// TIA Portal project "plc_main_V16" (V16)

(* hardware
DEVICE "S7-1200 station_1"  S7-1200 Station
   slot 0: "Rack_0"  S7-1200 Rack  Rack  V1.0
   slot 1: "PLC_main_ip_net_8"  CPU 1215C DC/DC/DC  6ES7 215-1AG40-0XB0  V4.2
DEVICE "PC-System_1"  SIMATIC PC station
   slot 0: "SIMATIC PC station"  Rail  SIMATIC PC-Station  V1.0
      slot 125: "Stationmanager"  Station_Manager  V6.0.4
   slot 1: "HMI_RT_1"  WinCC RT Advanced  6AV2 104-0xxxx-xxxx  16.0.0.0
      slot 33792: "Computer interface"  Host interface
   slot 2: "IE general_1"  IE General  IE_CP  V8.2.0
*)

// ===== PLC "PLC_main_ip_net_8"  CPU 1215C DC/DC/DC =====

VAR_GLOBAL   // PLC tag table "Default tag table"
   "Tag_1" AT %Q0.0 : Bool;
   "Tag_2" AT %Q0.1 : Bool;
   "LOGO_VM2" AT %MB100 : Byte;
   "LOGO_VM2.0" AT %M100.0 : Bool;
END_VAR

// folder: LGF/1 Date and timer operations/LGF_Astro

TYPE "LGF_typeAstroDMS"
VERSION : 0.1
   STRUCT
      dir : Char;   // Direction [N, S, E, W, n, s, e, w]
      deg : UInt;   // Degrees LAT [-89..+ 89]; LON [-179..+179]
      min : UInt;   // Minutes [0..+59]
      sec : UInt;   // Seconds [0..+59]
   END_STRUCT;
END_TYPE

// folder: LGF/8 Technology operations/LGF_NonLin

TYPE "LGF_typeNonLinSetpoints"
VERSION : 0.1
   STRUCT
      InputValue : Real;
      OutputValue : Real;
   END_STRUCT;
END_TYPE

// folder: LGF/8 Technology operations/LGF_Ramp

TYPE "LGF_typeRampTimeTable"
   STRUCT
      outVal : Real;
      "time" : Time;
   END_STRUCT;
END_TYPE

// folder: LGF/9 Measurement operations/LGF_RegressionLine

TYPE "LGF_typeRegressionLine"
   STRUCT
      x : Real;
      y : Real;
   END_STRUCT;
END_TYPE

// folder: Control_functions

DATA_BLOCK "control_DB"   // DB6
{ S7_Optimized_Access := 'FALSE' }
VERSION : 0.1
   VAR
      temperature_setpoint : Int;
      max_presure : Int := 40;
      emerg_coll_down : Bool;
      presure_err : Bool;
   END_VAR
BEGIN
END_DATA_BLOCK

DATA_BLOCK "LOGO"   // DB7
{ S7_Optimized_Access := 'FALSE' }
VERSION : 0.1
   VAR
      LOGO_heating_state : Bool;
   END_VAR
BEGIN
END_DATA_BLOCK

DATA_BLOCK "sensor_inputs"   // DB8
{ S7_Optimized_Access := 'TRUE' }
VERSION : 0.1
   VAR
      burning_temperature : Int;
      fire_state : Bool;
      flow_speed : Int;
      fluid_t : Int;
      system_presure : Int;
   END_VAR
BEGIN
END_DATA_BLOCK

DATA_BLOCK "actuators_output"   // DB9
{ S7_Optimized_Access := 'FALSE' }
VERSION : 0.1
   VAR
      gas_flow : Int;
      pimp_speed : Int;
      valve_state : Bool;
   END_VAR
BEGIN
END_DATA_BLOCK

DATA_BLOCK "Main_control_DB"   // DB10
{ S7_Optimized_Access := 'TRUE' }
VERSION : 0.1
// stored: InstanceOfName Main_control
"Main_control"
BEGIN
END_DATA_BLOCK

DATA_BLOCK "LGF_Impulse_DB_2"   // DB11
{ S7_Optimized_Access := 'TRUE' }
VERSION : 0.1
// stored: InstanceOfName LGF_Impulse
"LGF_Impulse"
BEGIN
END_DATA_BLOCK

// folder: Phisical_functions

DATA_BLOCK "phisical_DB"   // DB1
{ S7_Optimized_Access := 'TRUE' }
VERSION : 0.1
   VAR
      burning_t_old : Int;
      OUT_burning_t : Int;
      OUT_fire_state : Bool;
      OUT_fluid_t : Int;
      OUT_flow_speed : Int;
      IN_gas_flow : Int;
      IN_pimp_speed : Int;
      IN_valve_state : Bool;
      IN_pump_state : Bool;
      OUT_pump_err : Bool;
      OUT_pipe_err : Bool;
      OUT_tank_err : Bool;
      OUT_tank_presure : Int;
      OUT_residential_heeting : Bool;
      pump_failure : Bool := false;
      tank_failure : Bool := false;
      max_pump_failure_time : Time := T#10s;
      max_tank_presure : Int := 50;
   END_VAR
BEGIN
END_DATA_BLOCK

DATA_BLOCK "LGF_Impulse_DB"   // DB2
{ S7_Optimized_Access := 'TRUE' }
VERSION : 0.1
// stored: InstanceOfName LGF_Impulse
"LGF_Impulse"
BEGIN
END_DATA_BLOCK

DATA_BLOCK "LGF_Impulse_DB_1"   // DB3
{ S7_Optimized_Access := 'TRUE' }
VERSION : 0.1
// stored: InstanceOfName LGF_Impulse
"LGF_Impulse"
BEGIN
END_DATA_BLOCK

DATA_BLOCK "Phisical_proces_sim_dont_touch_DB_1"   // DB4
{ S7_Optimized_Access := 'TRUE' }
VERSION : 0.1
// stored: InstanceOfName Phisical_proces_sim_dont_touch
"Phisical_proces_sim_dont_touch"
BEGIN
END_DATA_BLOCK

// folder: System blocks/Program resources

DATA_BLOCK "IEC_Timer_0_DB"   // DB5
{ S7_Optimized_Access := 'TRUE' }
AUTHOR : Simatic
FAMILY : IEC
NAME : IEC_TMR
VERSION : 1.0
// stored: InstanceOfName IEC_TIMER
"IEC_TIMER"
BEGIN
END_DATA_BLOCK

// folder: (top level)

ORGANIZATION_BLOCK "Main"   // OB1, LAD, ProgramCycle
TITLE = "Main Program Sweep (Cycle)"
{ S7_Optimized_Access := 'TRUE' }
VERSION : 0.1
   VAR_INPUT
      Initial_Call : Bool;   // Initial call of this OB
      Remanence : Bool;   // =True, if remanent data are available
   END_VAR
BEGIN

REGION Network 1: Phisical proces
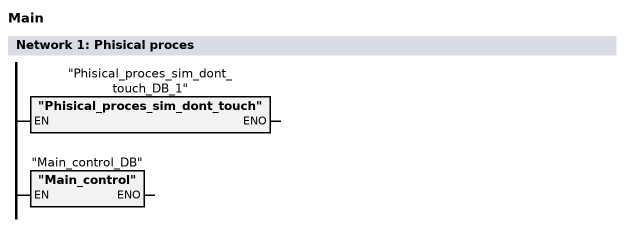
   RUNG wire#powerrail
      "Phisical_proces_sim_dont_touch_DB_1"()
   END_RUNG
   RUNG wire#powerrail
      "Main_control_DB"()
   END_RUNG
   // the same network as SCL:
   "Phisical_proces_sim_dont_touch_DB_1"();   // "Phisical_proces_sim_dont_touch"
   "Main_control_DB"();   // "Main_control"
END_REGION
END_ORGANIZATION_BLOCK

// folder: Control_functions

FUNCTION_BLOCK "Main_control"   // FB6, LAD
{ S7_Optimized_Access := 'TRUE' }
VERSION : 0.1
BEGIN

REGION Network 1
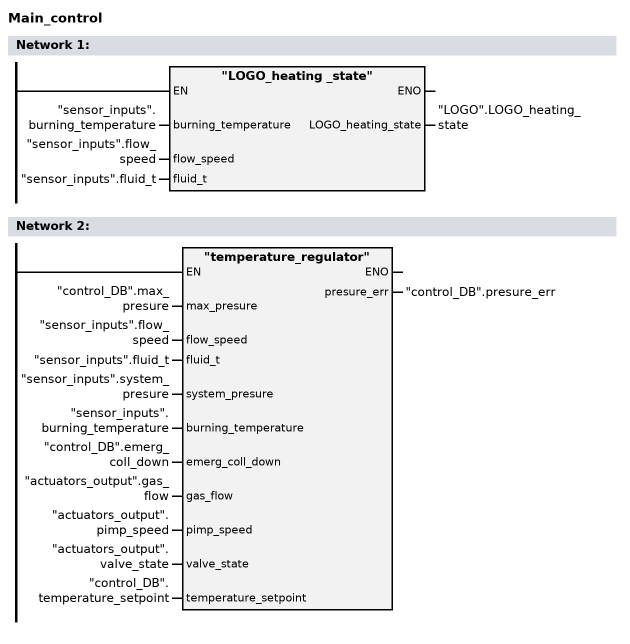
   RUNG wire#powerrail
      "LOGO_heating _state"(burning_temperature := "sensor_inputs".burning_temperature, flow_speed := "sensor_inputs".flow_speed, fluid_t := "sensor_inputs".fluid_t, LOGO_heating_state => "LOGO".LOGO_heating_state)
   END_RUNG
   // the same network as SCL:
   "LOGO_heating _state"(burning_temperature := "sensor_inputs".burning_temperature,
                         flow_speed := "sensor_inputs".flow_speed,
                         fluid_t := "sensor_inputs".fluid_t,
                         LOGO_heating_state => "LOGO".LOGO_heating_state);
END_REGION

REGION Network 2
   RUNG wire#powerrail
      "temperature_regulator"(max_presure := "control_DB".max_presure, flow_speed := "sensor_inputs".flow_speed, fluid_t := "sensor_inputs".fluid_t, system_presure := "sensor_inputs".system_presure, burning_temperature := "sensor_inputs".burning_temperature, emerg_coll_down := "control_DB".emerg_coll_down, gas_flow := "actuators_output".gas_flow, pimp_speed := "actuators_output".pimp_speed, valve_state := "actuators_output".valve_state, temperature_setpoint := "control_DB".temperature_setpoint, presure_err => "control_DB".presure_err)
   END_RUNG
   // the same network as SCL:
   "temperature_regulator"(max_presure := "control_DB".max_presure,
                           flow_speed := "sensor_inputs".flow_speed,
                           fluid_t := "sensor_inputs".fluid_t,
                           system_presure := "sensor_inputs".system_presure,
                           burning_temperature := "sensor_inputs".burning_temperature,
                           emerg_coll_down := "control_DB".emerg_coll_down,
                           gas_flow := "actuators_output".gas_flow,
                           pimp_speed := "actuators_output".pimp_speed,
                           valve_state := "actuators_output".valve_state,
                           temperature_setpoint := "control_DB".temperature_setpoint,
                           presure_err => "control_DB".presure_err);
END_REGION
END_FUNCTION_BLOCK

FUNCTION "LOGO_heating _state" : Void   // FC12, SCL
{ S7_Optimized_Access := 'TRUE' }
VERSION : 0.1
   VAR_INPUT
      burning_temperature : Int;
      flow_speed : Int;
      fluid_t : Int;
   END_VAR
   VAR_OUTPUT
      LOGO_heating_state : Bool;
   END_VAR
BEGIN
   IF #flow_speed > 1 AND #fluid_t > 15 THEN
       // Statement section IF
       #LOGO_heating_state := TRUE;
   ELSE
       #LOGO_heating_state := FALSE;
   END_IF;
END_FUNCTION

FUNCTION "temperature_regulator" : Void   // FC15, SCL
{ S7_Optimized_Access := 'TRUE' }
VERSION : 0.1
   VAR_INPUT
      max_presure : Int;
      flow_speed : Int;
      fluid_t : Int;
      system_presure : Int;
      burning_temperature : Int;
   END_VAR
   VAR_OUTPUT
      presure_err : Bool;
   END_VAR
   VAR_IN_OUT
      emerg_coll_down : Bool;
      gas_flow : Int;
      pimp_speed : Int;
      valve_state : Bool;
      temperature_setpoint : Int;
   END_VAR
   VAR_TEMP
      impulse : Bool;
   END_VAR
BEGIN
   "LGF_Impulse_DB_2"(frequency:=0.7,
                      impulse=>#impulse);

   IF #system_presure > #max_presure THEN
       // Statement section IF
       #temperature_setpoint := 0;
       #presure_err := true;
   END_IF;

   IF #impulse = TRUE THEN
       IF #temperature_setpoint > 0 THEN
           // Statement section IF
           #pimp_speed := 869;
       ELSE
           IF #pimp_speed > 0 THEN
               // Statement section IF
               #pimp_speed := #pimp_speed - 1;
           ELSE
               #pimp_speed := 0;
           END_IF;


       END_IF;
       // Statement section IF
       IF #temperature_setpoint > #fluid_t THEN
           // Statement section IF
           #gas_flow := #gas_flow + 1;
       ELSIF #temperature_setpoint < #fluid_t THEN
           #gas_flow := #gas_flow - 1;
       END_IF;

   END_IF;
END_FUNCTION

// folder: Phisical_functions

FUNCTION_BLOCK "Phisical_proces_sim_dont_touch"   // FB1, LAD
{ S7_Optimized_Access := 'TRUE' }
VERSION : 0.1
BEGIN

REGION Network 1
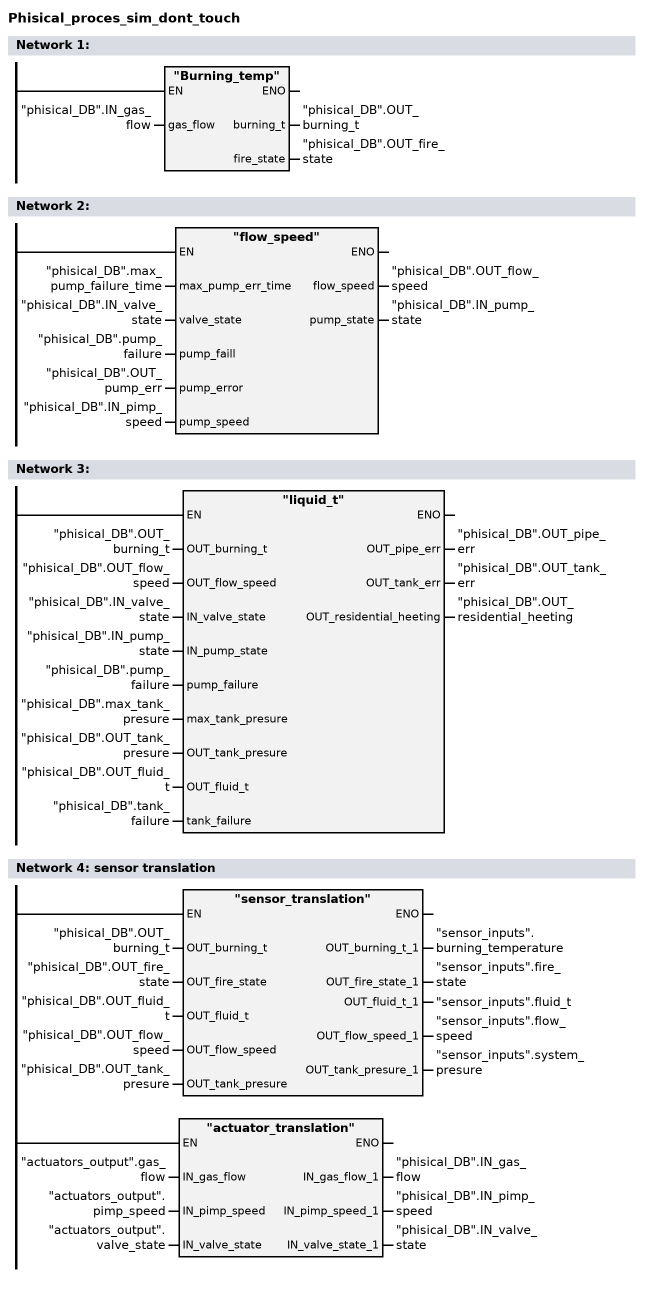
   RUNG wire#powerrail
      "Burning_temp"(gas_flow := "phisical_DB".IN_gas_flow, burning_t => "phisical_DB".OUT_burning_t, fire_state => "phisical_DB".OUT_fire_state)
   END_RUNG
   // the same network as SCL:
   "Burning_temp"(gas_flow := "phisical_DB".IN_gas_flow,
                  burning_t => "phisical_DB".OUT_burning_t,
                  fire_state => "phisical_DB".OUT_fire_state);
END_REGION

REGION Network 2
   RUNG wire#powerrail
      "flow_speed"(max_pump_err_time := "phisical_DB".max_pump_failure_time, valve_state := "phisical_DB".IN_valve_state, pump_faill := "phisical_DB".pump_failure, pump_error := "phisical_DB".OUT_pump_err, pump_speed := "phisical_DB".IN_pimp_speed, flow_speed => "phisical_DB".OUT_flow_speed, pump_state => "phisical_DB".IN_pump_state)
   END_RUNG
   // the same network as SCL:
   "flow_speed"(max_pump_err_time := "phisical_DB".max_pump_failure_time,
                valve_state := "phisical_DB".IN_valve_state,
                pump_faill := "phisical_DB".pump_failure,
                pump_error := "phisical_DB".OUT_pump_err,
                pump_speed := "phisical_DB".IN_pimp_speed,
                flow_speed => "phisical_DB".OUT_flow_speed,
                pump_state => "phisical_DB".IN_pump_state);
END_REGION

REGION Network 3
   RUNG wire#powerrail
      "liquid_t"(OUT_burning_t := "phisical_DB".OUT_burning_t, OUT_flow_speed := "phisical_DB".OUT_flow_speed, IN_valve_state := "phisical_DB".IN_valve_state, IN_pump_state := "phisical_DB".IN_pump_state, pump_failure := "phisical_DB".pump_failure, max_tank_presure := "phisical_DB".max_tank_presure, OUT_tank_presure := "phisical_DB".OUT_tank_presure, OUT_fluid_t := "phisical_DB".OUT_fluid_t, tank_failure := "phisical_DB".tank_failure, OUT_pipe_err => "phisical_DB".OUT_pipe_err, OUT_tank_err => "phisical_DB".OUT_tank_err, OUT_residential_heeting => "phisical_DB".OUT_residential_heeting)
   END_RUNG
   // the same network as SCL:
   "liquid_t"(OUT_burning_t := "phisical_DB".OUT_burning_t,
              OUT_flow_speed := "phisical_DB".OUT_flow_speed,
              IN_valve_state := "phisical_DB".IN_valve_state,
              IN_pump_state := "phisical_DB".IN_pump_state,
              pump_failure := "phisical_DB".pump_failure,
              max_tank_presure := "phisical_DB".max_tank_presure,
              OUT_tank_presure := "phisical_DB".OUT_tank_presure,
              OUT_fluid_t := "phisical_DB".OUT_fluid_t,
              tank_failure := "phisical_DB".tank_failure,
              OUT_pipe_err => "phisical_DB".OUT_pipe_err,
              OUT_tank_err => "phisical_DB".OUT_tank_err,
              OUT_residential_heeting => "phisical_DB".OUT_residential_heeting);
END_REGION

REGION Network 4: sensor translation
   RUNG wire#powerrail
      "sensor_translation"(OUT_burning_t := "phisical_DB".OUT_burning_t, OUT_fire_state := "phisical_DB".OUT_fire_state, OUT_fluid_t := "phisical_DB".OUT_fluid_t, OUT_flow_speed := "phisical_DB".OUT_flow_speed, OUT_tank_presure := "phisical_DB".OUT_tank_presure, OUT_burning_t_1 => "sensor_inputs".burning_temperature, OUT_fire_state_1 => "sensor_inputs".fire_state, OUT_fluid_t_1 => "sensor_inputs".fluid_t, OUT_flow_speed_1 => "sensor_inputs".flow_speed, OUT_tank_presure_1 => "sensor_inputs".system_presure)
   END_RUNG
   RUNG wire#powerrail
      "actuator_translation"(IN_gas_flow := "actuators_output".gas_flow, IN_pimp_speed := "actuators_output".pimp_speed, IN_valve_state := "actuators_output".valve_state, IN_gas_flow_1 => "phisical_DB".IN_gas_flow, IN_pimp_speed_1 => "phisical_DB".IN_pimp_speed, IN_valve_state_1 => "phisical_DB".IN_valve_state)
   END_RUNG
   // the same network as SCL:
   "sensor_translation"(OUT_burning_t := "phisical_DB".OUT_burning_t,
                        OUT_fire_state := "phisical_DB".OUT_fire_state,
                        OUT_fluid_t := "phisical_DB".OUT_fluid_t,
                        OUT_flow_speed := "phisical_DB".OUT_flow_speed,
                        OUT_tank_presure := "phisical_DB".OUT_tank_presure,
                        OUT_burning_t_1 => "sensor_inputs".burning_temperature,
                        OUT_fire_state_1 => "sensor_inputs".fire_state,
                        OUT_fluid_t_1 => "sensor_inputs".fluid_t,
                        OUT_flow_speed_1 => "sensor_inputs".flow_speed,
                        OUT_tank_presure_1 => "sensor_inputs".system_presure);
   "actuator_translation"(IN_gas_flow := "actuators_output".gas_flow,
                          IN_pimp_speed := "actuators_output".pimp_speed,
                          IN_valve_state := "actuators_output".valve_state,
                          IN_gas_flow_1 => "phisical_DB".IN_gas_flow,
                          IN_pimp_speed_1 => "phisical_DB".IN_pimp_speed,
                          IN_valve_state_1 => "phisical_DB".IN_valve_state);
END_REGION
END_FUNCTION_BLOCK

FUNCTION "Burning_temp" : Void   // FC1, SCL
{ S7_Optimized_Access := 'TRUE' }
VERSION : 0.1
   VAR_INPUT
      gas_flow : Int;
   END_VAR
   VAR_OUTPUT
      burning_t : Int;
      fire_state : Bool;
   END_VAR
   VAR_TEMP
      burning_t_temp : Int;
      triger : Bool;
   END_VAR
   VAR CONSTANT
      gas_to_temp : Int := 2;
   END_VAR
BEGIN
   //generates gas input state based on gas flow
   IF #gas_flow = 0 THEN
       #fire_state := FALSE;
   ELSE
       #fire_state := TRUE;
   END_IF;

   //Writing to phisicalDB
   #burning_t := #gas_flow * #gas_to_temp;
END_FUNCTION

FUNCTION "flow_speed" : Void   // FC10, SCL
{ S7_Optimized_Access := 'TRUE' }
VERSION : 0.1
   VAR_INPUT
      max_pump_err_time : Time;
      valve_state : Bool;
   END_VAR
   VAR_OUTPUT
      flow_speed : Int;
      pump_state : Bool;
   END_VAR
   VAR_IN_OUT
      pump_faill : Bool;
      pump_error : Bool;
      pump_speed : Int;
   END_VAR
   VAR_TEMP
      pump_err : Bool;
      impulse : Bool;
      countdown : Time;
      fault_timer_reset : Bool;
   END_VAR
   VAR CONSTANT
      rpm_to_l : Int := 10;
   END_VAR
BEGIN

   "LGF_Impulse_DB_1"(frequency:=70.0,
                      impulse=>#impulse,
                      countdown=>#countdown);

   IF #pump_faill = FALSE THEN
       // Statement section IF
       IF #pump_speed = 0 THEN
           // Statement section IF
           #pump_state := FALSE;
           #pump_err := FALSE;
       ELSE
           #pump_state := TRUE;

           IF #valve_state = FALSE THEN
               #flow_speed := 0;
               #pump_err := TRUE;
           ELSE

               #flow_speed := #pump_speed / #rpm_to_l;
               #pump_err := FALSE;

           END_IF;

       END_IF;
   ELSE
       #pump_state := TRUE;
       #pump_err := TRUE;
       #flow_speed := 0;
   END_IF;



       #pump_error := #pump_err;

       IF #pump_error = FALSE AND #pump_faill = FALSE THEN
           #fault_timer_reset := TRUE;
       ELSE
           #fault_timer_reset := FALSE;
       END_IF;

       "IEC_Timer_0_DB".TONR(IN:=#pump_error,
                             R:=#fault_timer_reset,
                             PT:=#max_pump_err_time,
                             Q=>#pump_faill
       );
END_FUNCTION

FUNCTION "liquid_t" : Void   // FC11, SCL
{ S7_Optimized_Access := 'TRUE' }
VERSION : 0.1
   VAR_INPUT
      OUT_burning_t : Int;
      OUT_flow_speed : Int;
      IN_valve_state : Bool;
      IN_pump_state : Bool;
      pump_failure : Bool;
      max_tank_presure : Int;
   END_VAR
   VAR_OUTPUT
      OUT_pipe_err : Bool;
      OUT_tank_err : Bool;
      OUT_residential_heeting : Bool;
   END_VAR
   VAR_IN_OUT
      OUT_tank_presure : Int;
      OUT_fluid_t : Int;
      tank_failure : Bool;
   END_VAR
   VAR_TEMP
      impulse : Bool;
      countdown : Time;
      valv_closes_increase : Int;
      pump_heat_decrease : Int;
      fluid_calculated_current : Int;
   END_VAR
   VAR CONSTANT
      fluid_to_burning_ratio : Int := 3;
   END_VAR
BEGIN
   "LGF_Impulse_DB"(frequency:=1.0,
                    impulse=>#impulse,
                    countdown=>#countdown);

   #valv_closes_increase := 0;

   #fluid_calculated_current := (#OUT_burning_t / #fluid_to_burning_ratio);

   (* IF #IN_valve_state = TRUE AND #IN_pump_state = TRUE THEN
       // Statement section IF
       #fluid_calculated_current := #fluid_calculated_current - #OUT_flow_speed / 8;
   END_IF; *)

   IF #impulse THEN


       (*
       HOW to create it so that when pump and valve doesnt work, temperature slowly increases
       *)

       IF #IN_valve_state = FALSE OR #IN_pump_state = FALSE OR #pump_failure = TRUE THEN

           IF #OUT_burning_t > #OUT_fluid_t THEN
               // Statement section IF
               #OUT_fluid_t := #OUT_fluid_t + 1;
           END_IF;

           IF #OUT_burning_t < #OUT_fluid_t THEN
               // Statement section IF
               #OUT_fluid_t := #OUT_fluid_t - 1;
           END_IF;

       ELSE
           IF #fluid_calculated_current > #OUT_fluid_t THEN
               // Statement section IF
               #OUT_fluid_t := #OUT_fluid_t + 1;
           END_IF;

           IF #fluid_calculated_current < #OUT_fluid_t THEN
               // Statement section IF
               #OUT_fluid_t := #OUT_fluid_t - 1;
           END_IF;
       END_IF;

       IF #tank_failure = TRUE THEN
           // Statement section IF
           #OUT_tank_presure := #OUT_tank_presure - 5;
       ELSE
           #OUT_tank_presure := ((#OUT_fluid_t) / 2.83);
       END_IF;
   END_IF;





   IF #tank_failure = FALSE THEN
       IF #OUT_tank_presure > #max_tank_presure THEN
           #tank_failure := TRUE;
       END_IF;
   END_IF;



   IF #OUT_fluid_t > 30 & #IN_valve_state = TRUE & #IN_pump_state = TRUE THEN
       IF #pump_failure = TRUE THEN

           #OUT_residential_heeting := FALSE;
       ELSE
           #OUT_residential_heeting := TRUE;
       END_IF;


   ELSE
       #OUT_residential_heeting := FALSE;
   END_IF;
END_FUNCTION

FUNCTION "sensor_translation" : Void   // FC13, SCL
{ S7_Optimized_Access := 'TRUE' }
VERSION : 0.1
   VAR_INPUT
      OUT_burning_t : Int;
      OUT_fire_state : Bool;
      OUT_fluid_t : Int;
      OUT_flow_speed : Int;
      OUT_tank_presure : Int;
   END_VAR
   VAR_OUTPUT
      OUT_burning_t_1 : Int;
      OUT_fire_state_1 : Bool;
      OUT_fluid_t_1 : Int;
      OUT_flow_speed_1 : Int;
      OUT_tank_presure_1 : Int;
   END_VAR
BEGIN
   #OUT_burning_t_1 := #OUT_burning_t;
   #OUT_fire_state_1 := #OUT_fire_state;
   #OUT_fluid_t_1 := #OUT_fluid_t;
   #OUT_flow_speed_1 := #OUT_flow_speed;
   #OUT_tank_presure_1 := #OUT_tank_presure;
END_FUNCTION

FUNCTION "actuator_translation" : Void   // FC14, SCL
{ S7_Optimized_Access := 'TRUE' }
VERSION : 0.1
   VAR_INPUT
      IN_gas_flow : Int;
      IN_pimp_speed : Int;
      IN_valve_state : Bool;
   END_VAR
   VAR_OUTPUT
      IN_gas_flow_1 : Int;
      IN_pimp_speed_1 : Int;
      IN_valve_state_1 : Bool;
   END_VAR
BEGIN
   #IN_gas_flow_1 := #IN_gas_flow;
   #IN_pimp_speed_1 := #IN_pimp_speed;
   #IN_valve_state_1 := #IN_valve_state;
END_FUNCTION

// folder: Phisical_functions/LGF/0 Bit logic operations

FUNCTION_BLOCK "LGF_PulseRelay"   // FB3, SCL
{ S7_Optimized_Access := 'TRUE' }
VERSION : 0.1
   VAR_INPUT
      trigger : Bool;   // trigger signal, rising edge
      set : Bool;   // set signal. rising edge
      reset : Bool;   // reset signal, rising edge
   END_VAR
   VAR_OUTPUT
      out : Bool;   // output signal
   END_VAR
   VAR
      statTriggerOld : Bool := false;   // -
      statTriggerRis : Bool := false;   // -
      statSetOld : Bool := false;   // -
      statSetRis : Bool := false;   // -
      statResetOld : Bool := false;   // -
      statResetRis : Bool := false;   // -
      statOut : Bool := false;   // -
   END_VAR
BEGIN
   //=============================================================================
   // SIEMENS AG
   // (c)Copyright 2017 
   //-----------------------------------------------------------------------------
   // Library:       LGF (Library General Functions)
   // Tested with:   CPU1212C DC/DC/DC FW:V4.2
   // Engineering:   TIA Portal V14 Update 1
   // Restrictions:  -
   // Requirements:  PLC (S7-1200 / S7-1500)
   // Functionality: Pulse relay, Surge relay, Toggle-Flip-Flop, Frequency divider
   //-----------------------------------------------------------------------------
   // Change log table:
   // Version Date        In charge / Changes applied
   // 01.00.00 06.06.2015 Siemens Industry Online Support
   //                     First released version
   // 01.00.01 02.01.2017 Siemens Industry Online Support
   //                     Upgrade: TIA V14 Update 1
   // 01.00.02 02.01.2017 Siemens Industry Online Support
   //                     Comment correction                  
   // 01.00.03 17.08.2018 Siemens Industry Online Support
   //                     Upgrade: TIA V15 Update 2
   // 01.00.04 23.11.2018 Siemens Industry Online Support
   //                     Upgrade: TIA V15.1
   //=============================================================================

   // Scan for risign edge "trigger"
   IF #trigger AND  NOT #statTriggerOld THEN
     #statTriggerRis := TRUE;
   ELSE
     #statTriggerRis := FALSE;
   END_IF;
   #statTriggerOld := #trigger;

   // Scan for risign edge "set"
   IF #set AND NOT #statSetOld THEN
     #statSetRis := TRUE;
   ELSE
     #statSetRis := FALSE;
   END_IF;
   #statSetOld := #set;

   // Scan for risign edge "reset"
   IF #reset AND NOT #statResetOld THEN
     #statResetRis := TRUE;
   ELSE
     #statResetRis := FALSE;
   END_IF;
   #statResetOld := #reset;

   // Create toggle signal
   IF #statTriggerRis AND NOT #statOut THEN
     #statOut := TRUE;
   ELSIF #statTriggerRis AND #statOut THEN
     #statOut := FALSE;
   END_IF;

   // Output: toggle, set, reset
   IF #statTriggerRis THEN
     #out := #statOut;
   END_IF;

   IF #statSetRis THEN
     #out := TRUE;
   END_IF;

   IF #statResetRis THEN
     #out := FALSE;
   END_IF;
END_FUNCTION_BLOCK

// folder: Phisical_functions/LGF/1 Date and timer operations

FUNCTION_BLOCK "LGF_SetTime"   // FB4, SCL
{ S7_Optimized_Access := 'TRUE' }
VERSION : 0.1
   VAR_INPUT
      setSystemTimeUTC : Bool;   // Set system time
      systemTimeUTC : DTL;   // System time
      setLocalTime : Bool;   // Set local time
      localTime : DTL;   // Local Time
      setTimeZone : Bool;   // Set time zone and daylight saving time
      timeZone : Int;   // Timezones HHMM [-1200.. -330.. 0.. 930.. 1200.. 1300]
      daylightSavingTime : Bool;   // Daylight saving time: activated [1], deactivated [0]
   END_VAR
   VAR_OUTPUT
      actSystemTime : DTL;   // -
      actLocalTime : DTL;   // -
      lastSetTimeZone : String;   // Time zone that was set last by this block
      error : Bool;   // Error
      status : Word;   // Status and error codes
      statusID : UInt;   // Error destination: "1" = LGF_SetTime; "2" = SET_TIMEZONE
   END_VAR
   VAR
      statSetSystemTimeOld : Bool;   // -
      statSetLocalTimeOld : Bool;   // -
      statSetTimeZoneOld : Bool;   // -
      statTimeZone : TimeTransformationRule;   // -
      InstSET_TIMEZONE : SET_TIMEZONE;   // -
   END_VAR
   VAR_TEMP
      tempSetLocalTimeRet : Int;   // -
      tempSetSystemTimeRet : Int;   // -
      tempSystemTimeRet : Int;   // -
      tempLocalTimeRet : Int;   // -
      tempTimeZoneDone : Bool;   // -
      tempTimeZoneBusy : Bool;   // -
      tempTimeZoneError : Bool;   // -
      tempTimeZoneStatus : Word;   // -
   END_VAR
   VAR CONSTANT
      HOUR : Int := 60;   // -
      "30MIN" : Int := 30;   // -
      "15MIN" : Int := 15;   // -
      "0MIN" : Int := 0;   // -
      NO_ERROR : Word := 16#0000;   // -
      NO_CURRENT_JOBS : Word := 16#7000;   // -
      ERROR_NO_DEFINED_TIME_ZONE : Word := 16#8200;   // No defined time zone is selected; check input "timeZone"
      ERROR_IN_THIS_BLOCK : UInt := 1;   // Error in this block
      ERROR_SET_TIMEZONE : UInt := 2;   // Error instruction SET_TIMEZONE
   END_VAR
   // statTimeZone.Bias := 0;
   // statTimeZone.DaylightBias := 60;
   // statTimeZone.DaylightStartMonth := 3;
   // statTimeZone.DaylightStartWeek := 5;
   // statTimeZone.DaylightStartWeekday := 1;
   // statTimeZone.DaylightStartHour := 2;
   // statTimeZone.DaylightStartMinute := 0;
   // statTimeZone.StandardStartMonth := 10;
   // statTimeZone.StandardStartWeek := 5;
   // statTimeZone.StandardStartWeekday := 1;
   // statTimeZone.StandardStartHour := 3;
   // statTimeZone.StandardStartMinute := 0;
   // statTimeZone.TimeZoneName := 'not even set by LGF_TimeZone';
BEGIN
   //=============================================================================
   // SIEMENS AG
   // (c)Copyright 2017 
   //-----------------------------------------------------------------------------
   // Library:       LGF (Library General Functions)
   // Tested with:   CPU1212C DC/DC/DC FW:V4.2
   // Engineering:   TIA Portal V14 Update 1
   // Restrictions:  -
   // Requirements:  PLC (S7-1200 / S7-1500)
   // Functionality: Set system time, local time, time zone
   //-----------------------------------------------------------------------------
   // Change log table:
   // Version Date         In charge / Changes applied
   // 01.00.00 08.06.2015  Siemens Industry Online Support
   //                      First released version
   // 01.00.01 02.01.2017  Siemens Industry Online Support
   //                      Upgrade: TIA V14 Update 1
   // 01.00.02 02.03.2017  Siemens Industry Online Support
   //                      Bugfix: FB number: automatic
   // 01.00.03 17.08.2018  Siemens Industry Online Support
   //                      Upgrade: TIA V15 Update 2
   // 01.00.04 23.11.2018  Siemens Industry Online Support
   //                      Upgrade: TIA V15.1
   // 01.00.05 20.02.2019  Siemens Industry Online Support
   //                      Bugfix: Rising edge at input REQ of SET_TIMEOUT
   // =============================================================================

   // Set "No current job" status
   #error := false;
   #statusID := #ERROR_IN_THIS_BLOCK;
   #status := #NO_CURRENT_JOBS;

   // Reading system and local time
   #tempSystemTimeRet := RD_SYS_T(#actSystemTime); // Output current system time
   #tempLocalTimeRet := RD_LOC_T(#actLocalTime); // Output current local

   // Set system time by rising edge =============================================
   IF #setSystemTimeUTC AND NOT #statSetSystemTimeOld THEN
     #tempSetSystemTimeRet := WR_SYS_T(#systemTimeUTC);
   END_IF;
   #statSetSystemTimeOld := #setSystemTimeUTC;

   // Set local time zone by rising edge =========================================
   IF #setLocalTime AND NOT #statSetLocalTimeOld THEN
     #tempSetLocalTimeRet := WR_LOC_T(LOCTIME := #localTime, DST := #daylightSavingTime);
   END_IF;
   #statSetLocalTimeOld := #setLocalTime;

   // Set time zone by rising edge ===============================================
   IF #setTimeZone AND NOT #statSetTimeZoneOld THEN
     CASE #timeZone OF
       -1200:  // (UTC -12:00) Eniwetok, Kwajalein
         #statTimeZone.Bias := -12 * #HOUR;
         #statTimeZone.TimeZoneName := '(UTC -12:00)';
       -1100:  // (UTC -11:00) Midway Island
         #statTimeZone.Bias := -11 * #HOUR;
         #statTimeZone.TimeZoneName := '(UTC -11:00)';
       -1000:  // (UTC -10:00) Hawaii
         #statTimeZone.Bias := -10 * #HOUR;
         #statTimeZone.TimeZoneName := '(UTC -10:00)';
       -930:  // (UTC -09:30) (French) Polynesia
         #statTimeZone.Bias := -9 * #HOUR + #"30MIN";
         #statTimeZone.TimeZoneName := '(UTC -09:00)';
       -900:  // (UTC -09:00) Alaska
         #statTimeZone.Bias := -9 * #HOUR;
         #statTimeZone.TimeZoneName := '(UTC -09:00)';
       -800:  // (UTC -08:00) Tijuana, Los Angeles, Seattle, Vancouver
         #statTimeZone.Bias := -8 * #HOUR;
         #statTimeZone.TimeZoneName := '(UTC -08:00)';
       -700:  // (UTC -07:00) Arizona, Denver, Salt Lake City, Calgary
         #statTimeZone.Bias := -7 * #HOUR;
         #statTimeZone.TimeZoneName := '(UTC -07:00)';
       -600:  // (UTC -06:00) Chicago, Dallas, Kansas City, Winnipeg
         #statTimeZone.Bias := -6 * #HOUR;
         #statTimeZone.TimeZoneName := '(UTC -06:00)';
       -500:  // (UTC -05:00) Eastern Time (USA & Canada)
         #statTimeZone.Bias := -5 * #HOUR;
         #statTimeZone.TimeZoneName := '(UTC -05:00)';
       -400:  // (UTC -04:00) La Paz, Georgetown
         #statTimeZone.Bias := -4 * #HOUR;
         #statTimeZone.TimeZoneName := '(UTC -04:00)';
       -330:  // (UTC -03:30) Newfoundland
         #statTimeZone.Bias := -3 * #HOUR + #"30MIN";
         #statTimeZone.TimeZoneName := '(UTC -03:30)';
       -300:  // (UTC -03:00) Brasilia, Buenos Aires
         #statTimeZone.Bias := -3 * #HOUR;
         #statTimeZone.TimeZoneName := '(UTC -03:00)';
       -200:  // (UTC -02:00) Mid-Atlantic
         #statTimeZone.Bias := -2 * #HOUR;
         #statTimeZone.TimeZoneName := '(UTC -02:00)';
       -100:  // (UTC -01:00) Azores, Cape Verde Is.
         #statTimeZone.Bias := -1 * #HOUR;
         #statTimeZone.TimeZoneName := '(UTC -01:00)';
       0:  // (UTC) Dublin, Edinburgh, Lisbon, London
         #statTimeZone.Bias := 0;
         #statTimeZone.TimeZoneName := '(UTC)';
       100:  // (UTC +01:00) Berlin, Bern, Brussels, Rome, Stockholm, Vienna
         #statTimeZone.Bias := 1 * #HOUR;
         #statTimeZone.TimeZoneName := '(UTC +01:00)';
       200: // (UTC +02:00) Athens, Istanbul, Minsk, Bucharest
         #statTimeZone.Bias := 2 * #HOUR;
         #statTimeZone.TimeZoneName := '(UTC +02:00)';
       300: // (UTC +03:00) Baghdad, Kuwait, Riyadh
         #statTimeZone.Bias := 3 * #HOUR;
         #statTimeZone.TimeZoneName := '(UTC +03:00)';
       330: // (UTC +03:00) Iran
         #statTimeZone.Bias := 3 * #HOUR + #"30MIN";
         #statTimeZone.TimeZoneName := '(UTC +03:30)';
       400: // (UTC +04:00) Moscow, St. Petersburg, Volgograd, Abu Dhabi, Muscat
         #statTimeZone.Bias := 4 * #HOUR;
         #statTimeZone.TimeZoneName := '(UTC +04:00)';
       430: // (UTC +04:30) Afghanistan
         #statTimeZone.Bias := 4 * #HOUR + #"30MIN";
         #statTimeZone.TimeZoneName := '(UTC +04:30)';
       500: // (UTC +05:00) Islamabad, Karachi, Tashkent
         #statTimeZone.Bias := 5 * #HOUR;
         #statTimeZone.TimeZoneName := '(UTC +05:00)';
       530: // (UTC +05:30) India, Sri Lanka
         #statTimeZone.Bias := 5 * #HOUR + #"30MIN";
         #statTimeZone.TimeZoneName := '(UTC +05:30)';
       545: // (UTC +05:45) India, Sri Lanka
         #statTimeZone.Bias := 5 * #HOUR + #"30MIN" + #"15MIN";
         #statTimeZone.TimeZoneName := '(UTC +05:45)';
       600: // (UTC +06:00) Astana, Almaty, Dhaka, Colombo
         #statTimeZone.Bias := 6 * #HOUR;
         #statTimeZone.TimeZoneName := '(UTC +06:00)';
       630: // (UTC +06:30) Coco Island, Mayanmar
         #statTimeZone.Bias := 6 * #HOUR + #"30MIN";
         #statTimeZone.TimeZoneName := '(UTC +06:30)';
       700: // (UTC +07:00) Bangkok, Hanoi, Jakarta
         #statTimeZone.Bias := 7 * #HOUR;
         #statTimeZone.TimeZoneName := '(UTC +07:00)';
       800: // (UTC +08:00) Beijing, Chongqing, Hong Kong, Urumqi
         #statTimeZone.Bias := 8 * #HOUR;
         #statTimeZone.TimeZoneName := '(UTC +08:00)';
       830: // (UTC +08:30) North Corea
         #statTimeZone.Bias := 8 * #HOUR + #"30MIN";
         #statTimeZone.TimeZoneName := '(UTC +08:30)';
       900: // (UTC +09:00) Yakutsk, Osaka, Sapporo, Tokyo, Seoul
         #statTimeZone.Bias := 9 * #HOUR;
         #statTimeZone.TimeZoneName := '(UTC +09:00)';
       930: // (UTC +09:30) Australia: Northern Territory, South Australia
         #statTimeZone.Bias := 9 * #HOUR + #"30MIN";
         #statTimeZone.TimeZoneName := '(UTC +09:30)';
       1000: // (UTC +10:00) Brisbane, Canberra, Melbourne, Sydney
         #statTimeZone.Bias := 10 * #HOUR;
         #statTimeZone.TimeZoneName := '(UTC +10:00)';
       1030: // (UTC +10:30) Australia: Lord Howe Island
         #statTimeZone.Bias := 10 * #HOUR + #"30MIN";
         #statTimeZone.TimeZoneName := '(UTC +10:30)';
       1100: // (UTC +11:00) Vladivostok, Magadan, Solomon Is., New Caledonia
         #statTimeZone.Bias := 11 * #HOUR;
         #statTimeZone.TimeZoneName := '(UTC +11:00)';
       1200: // (UTC +12:00) Auckland, Wellington
         #statTimeZone.Bias := 12 * #HOUR;
         #statTimeZone.TimeZoneName := '(UTC +12:00)';
       1245: // (UTC +12:45) Chatham Islands
         #statTimeZone.Bias := 12 * #HOUR + #"30MIN" + #"15MIN";
         #statTimeZone.TimeZoneName := '(UTC +12:45)';
       1300: // (UTC +13:00) Kiribati
         #statTimeZone.Bias := 13 * #HOUR;
         #statTimeZone.TimeZoneName := '(UTC +13:00)';
       ELSE  // Error handling
         #error := true;
         #statusID := #ERROR_IN_THIS_BLOCK;
         #status := #ERROR_NO_DEFINED_TIME_ZONE;
         RETURN;
     END_CASE;
   END_IF;

   // Select daylight saving time on/off
   IF #daylightSavingTime THEN
     #statTimeZone.DaylightBias := #HOUR;
   ELSE
     #statTimeZone.DaylightBias := #"0MIN";
   END_IF;

   // Set time zone by rising edge (REQ)
   #InstSET_TIMEZONE(REQ := (#setTimeZone AND NOT #statSetTimeZoneOld),
                     TimeZone := #statTimeZone,
                     DONE => #tempTimeZoneDone,
                     BUSY => #tempTimeZoneBusy,
                     ERROR => #tempTimeZoneError,
                     STATUS => #tempTimeZoneStatus);

   #statSetTimeZoneOld := #setTimeZone;

   IF #tempTimeZoneError THEN
     #error := true;
     #statusID := #ERROR_SET_TIMEZONE;
     #status := #tempTimeZoneStatus;
     RETURN;
   END_IF;

   // Output the last set time zone
   #lastSetTimeZone := #statTimeZone.TimeZoneName;

   // No errors
   #status := #NO_ERROR;
END_FUNCTION_BLOCK

FUNCTION_BLOCK "LGF_TimerSwitch"   // FB10002, SCL
{ S7_Optimized_Access := 'TRUE' }
   VAR_INPUT
      onMonth : USInt;   // Month, in which the signal shall be set.
      onDay : USInt;   // Day, at which the signal shall be set.
      onWeekday : USInt;   // Sunday: 1, Monday: 2, Tuesday: 3, ...
      onHour : USInt;   // Hour, at which the signal shall be set.
      onMinute : USInt;   // Minute, at which the signal shall be set.
      offMonth : USInt;   // Month, in which the signal shall be reset.
      offDay : USInt;   // Day, at which the signal shall be reset.
      offWeekday : USInt;   // Sunday: 1, Monday: 2, Tuesday: 3, ...
      offHour : USInt;   // Hour, at which the signal shall be reset.
      offMinute : USInt;   // Minute, at which the signal shall be reset.
      mode : USInt;   // Daily: 1, weekly: 2, monthly: 3, yearly: 4, workday: 5, weekend: 6
   END_VAR
   VAR_OUTPUT
      signal : Bool;   // Output signal
      actLocalTime : DTL;   // Current local time
      error : Bool;   // "0" = no error; "1" = error
      statusID : UInt;   // Error destination: "1" = LGF_TimerSwitch; "2" = RD_LOC_T
      status : Word;   // Status and error codes
   END_VAR
   VAR_TEMP
      tempSignal : Bool;   // -
      tempTime : DTL;   // -
      tempReadTimeStatus : Int;   // -
      tempOnTime : DTL;   // -
      tempOnTimeTOD : Time_Of_Day;   // -
      tempOffTime : DTL;   // -
      tempOffTimeTOD : Time_Of_Day;   // -
      tempActTime : DTL;   // -
      tempActTimeTOD : Time_Of_Day;   // -
      tempCrossMidnight : Bool;   // -
   END_VAR
   VAR CONSTANT
      NO_ERROR : Word := 16#0000;   // -
      NO_CURRENT_JOBS : Word := 16#7000;   // -
      NO_MODE_SELECTED : Word := 16#8200;   // No suitable mode is selected, check input "mode"
      ERROR_IN_THIS_BLOCK : UInt := 1;   // Error in this block
      ERROR_RD_LOC_T : UInt := 2;   // Error in function RD_LOC_T
   END_VAR
BEGIN
   //=============================================================================
   // SIEMENS AG
   // (c)Copyright 2017
   //-----------------------------------------------------------------------------
   // Library:       LGF (Library General Functions)
   // Tested with:   CPU1212C DC/DC/DC FW:V4.2
   // Engineering:   TIA Portal V14 Update 1
   // Restrictions:  -
   // Requirements:  PLC (S7-1200 / S7-1500)
   // Functionality: Timer Switch (daily, weekly, monthly, working days, ...)
   //-----------------------------------------------------------------------------
   // Change log table:
   // Version Date         In charge / Changes applied
   // 01.00.00 19.08.2015  Siemens Industry Online Support
   //                      First released version
   // 01.00.01 16.11.2015  Siemens Industry Online Support
   //                      Fix in mode 2
   // 01.01.00 23.05.2016  Siemens Industry Online Support
   //                      New mode 5 + 6
   //                      New output: actLocalTime
   // 01.01.01 02.01.2017  Siemens Industry Online Support
   //                      Upgrade: TIA V14 Update 1
   // 01.01.02 14.09.2018  Siemens Industry Online Support
   //                      Fix in modes 1, 3, 5, 6                    
   // 01.01.03 17.09.2018  Siemens Industry Online Support
   //                      Upgrade: TIA V15 Update 2
   // 01.01.04 10.10.2018  Siemens Industry Online Support
   //                      Connection to type restored
   // 01.01.05 23.11.2018  Siemens Industry Online Support
   //                      Upgrade: TIA V15.1
   //=============================================================================

   //Set "No current job" status
   #error := false;
   #statusID := #ERROR_IN_THIS_BLOCK;
   #status := #NO_CURRENT_JOBS;

   //Read local time
   #tempReadTimeStatus := RD_LOC_T(#tempTime);
   #actLocalTime := #tempTime;

   IF (#tempReadTimeStatus > 1)
   THEN
     #error := true;
     #statusID := #ERROR_RD_LOC_T;
     #status := INT_TO_WORD(#tempReadTimeStatus);
     RETURN;
   END_IF;


   #tempOnTime.HOUR := #onHour;
   #tempOnTime.MINUTE := #onMinute;
   #tempOnTime.SECOND := 0;
   #tempOnTime.NANOSECOND := 0;

   #tempOffTime.HOUR := #offHour;
   #tempOffTime.MINUTE := #offMinute;
   #tempOffTime.SECOND := 0;
   #tempOffTime.NANOSECOND := 0;

   CASE #mode OF
     1:  // Mode: daily
       #tempOnTime.YEAR := #tempTime.YEAR;
       #tempOnTime.MONTH := #tempTime.MONTH;
       #tempOnTime.WEEKDAY := #tempTime.WEEKDAY;
       #tempOnTime.DAY := #tempTime.DAY;

       #tempOnTimeTOD := DTL_TO_TOD(#tempOnTime);

       #tempOffTime.YEAR := #tempTime.YEAR;
       #tempOffTime.MONTH := #tempTime.MONTH;
       #tempOffTime.WEEKDAY := #tempTime.WEEKDAY;
       #tempOffTime.DAY := #tempTime.DAY;

       #tempOffTimeTOD := DTL_TO_TOD(#tempOffTime);
       #tempActTimeTOD := DTL_TO_TOD(#tempTime);

       IF (#tempOnTimeTOD > #tempOffTimeTOD)
       THEN
         IF (#tempActTimeTOD > #tempOffTimeTOD)
         THEN
           #tempOffTime := #tempOffTime + t#1d;
         ELSE
           #tempOnTime := #tempOnTime - t#1d;
         END_IF;
       END_IF;

       IF (#tempTime >= #tempOnTime)
         AND (#tempTime < #tempOffTime)
       THEN
         #tempSignal := true;
       ELSE
         #tempSignal := false;
       END_IF;

       #signal := #tempSignal;

     2:  // Mode: weekly
       #tempOnTime.YEAR := 2015;
       #tempOnTime.MONTH := 1;
       #tempOnTime.DAY := #onWeekday + 3;

       #tempOnTimeTOD := DTL_TO_TOD(#tempOnTime);

       #tempOffTime.YEAR := 2015;
       #tempOffTime.MONTH := 1;
       #tempOffTime.DAY := #offWeekday + 3;

       #tempOffTimeTOD := DTL_TO_TOD(#tempOffTime);

       #tempActTime := #tempTime;
       #tempActTime.YEAR := 2015;
       #tempActTime.MONTH := 1;
       #tempActTime.DAY := #tempActTime.WEEKDAY + 3;

       #tempActTimeTOD := DTL_TO_TOD(#tempTime);

       IF (#onWeekday > #offWeekday)
         OR ((#onWeekday = #offWeekday)
         AND (#tempOnTimeTOD > #tempOffTimeTOD))
       THEN
         #tempOffTime.DAY := #offWeekday + 10;
         IF (#tempActTime.WEEKDAY < #onWeekday)
           OR ((#onWeekday = #offWeekday)
           AND (#tempActTimeTOD < #tempOffTimeTOD))
         THEN
           #tempActTime.DAY := #tempActTime.WEEKDAY + 10;
         END_IF;
       END_IF;

       IF (#tempActTime >= #tempOnTime)
         AND (#tempActTime < #tempOffTime)
       THEN
         #tempSignal := true;
       ELSE
         #tempSignal := false;
       END_IF;

       #signal := #tempSignal;

     3:  // Mode: monthly
       #tempOnTime.YEAR := #tempTime.YEAR;
       #tempOnTime.MONTH := #tempTime.MONTH;
       #tempOnTime.WEEKDAY := #tempTime.WEEKDAY;
       #tempOnTime.DAY := #onDay;

       #tempOnTimeTOD := DTL_TO_TOD(#tempOnTime);

       #tempOffTime.YEAR := #tempTime.YEAR;
       #tempOffTime.MONTH := #tempTime.MONTH;
       #tempOffTime.WEEKDAY := #tempTime.WEEKDAY;
       #tempOffTime.DAY := #offDay;

       #tempOffTimeTOD := DTL_TO_TOD(#tempOffTime);
       #tempActTimeTOD := DTL_TO_TOD(#tempTime);

       IF (#onDay > #offDay)
         OR ((#onDay = #offDay)
         AND (#tempOnTimeTOD > #tempOffTimeTOD))
       THEN
         IF (#tempTime.DAY > #offDay)
           OR ((#tempTime.DAY = #offDay)
           AND (#tempActTimeTOD > #tempOffTimeTOD))
         THEN
           #tempOffTime.MONTH := #tempOffTime.MONTH + 1;

           IF (#tempOffTime.MONTH > 12)
           THEN
             #tempOffTime.MONTH := 1;
             #tempOffTime.YEAR := #tempOffTime.YEAR + 1;
           END_IF;

         ELSE
           #tempOnTime.MONTH := #tempOnTime.MONTH - 1;

           IF (#tempOnTime.MONTH < 1)
           THEN
             #tempOnTime.MONTH := 12;
             #tempOnTime.YEAR := #tempOnTime.YEAR - 1;
           END_IF;

         END_IF;
       END_IF;


       IF (#tempTime >= #tempOnTime)
         AND (#tempTime < #tempOffTime)
       THEN
         #tempSignal := true;
       ELSE
         #tempSignal := false;
       END_IF;

       #signal := #tempSignal;

     4:  // Mode: yearly
       #tempOnTime.YEAR := #tempTime.YEAR;
       #tempOnTime.MONTH := #onMonth;
       #tempOnTime.WEEKDAY := #tempTime.WEEKDAY;
       #tempOnTime.DAY := #onDay;

       #tempOnTimeTOD := DTL_TO_TOD(#tempOnTime);

       #tempOffTime.YEAR := #tempTime.YEAR;
       #tempOffTime.MONTH := #offMonth;
       #tempOffTime.WEEKDAY := #tempTime.WEEKDAY;
       #tempOffTime.DAY := #offDay;

       #tempOffTimeTOD := DTL_TO_TOD(#tempOffTime);
       #tempActTimeTOD := DTL_TO_TOD(#tempTime);

       IF (#onMonth > #offMonth)
         OR ((#onMonth = #offMonth)
         AND (#tempOnTimeTOD > #tempOffTimeTOD))
       THEN
         IF (#tempTime.MONTH > #offMonth)
           OR ((#tempTime.MONTH = #offMonth)
           AND (#tempActTimeTOD > #tempOffTimeTOD))
         THEN
           #tempOffTime.YEAR := #tempOffTime.YEAR + 1;
         ELSE
           #tempOnTime.YEAR := #tempOnTime.YEAR - 1;
         END_IF;
       END_IF;

       IF (#tempTime >= #tempOnTime)
         AND (#tempTime < #tempOffTime)
       THEN
         #tempSignal := true;
       ELSE
         #tempSignal := false;
       END_IF;

       #signal := #tempSignal;

     5:  // Mode: working days (Monday - Friday)    
       #tempOnTime.YEAR := 2015;
       #tempOnTime.MONTH := 1;
       #tempOnTime.DAY := #tempTime.WEEKDAY + 3;

       #tempOnTimeTOD := DTL_TO_TOD(#tempOnTime);

       #tempOffTime.YEAR := 2015;
       #tempOffTime.MONTH := 1;
       #tempOffTime.DAY := #tempTime.WEEKDAY + 3;

       #tempOffTimeTOD := DTL_TO_TOD(#tempOffTime);

       #tempActTime := #tempTime;
       #tempActTime.YEAR := 2015;
       #tempActTime.MONTH := 1;
       #tempActTime.DAY := #tempActTime.WEEKDAY + 3;

       #tempActTimeTOD := DTL_TO_TOD(#tempTime);

       IF (#tempOnTimeTOD > #tempOffTimeTOD)
       THEN
         #tempCrossMidnight := TRUE;
         IF (#tempActTimeTOD > #tempOffTimeTOD)
         THEN
           #tempOffTime := #tempOffTime + t#1d;
         ELSE
           #tempOnTime := #tempOnTime - t#1d;
         END_IF;
       ELSE
         #tempCrossMidnight := FALSE;
       END_IF;

       IF (#tempOnTime.DAY <= 5)
       THEN
         #tempOnTime.DAY := 5;
       ELSIF (#tempOnTime.DAY > 9)
       THEN
         #tempOnTime.DAY := 9;
       END_IF;

       IF (#tempOffTime.DAY > 9)
         AND (#tempCrossMidnight = TRUE)
       THEN
         #tempOffTime.DAY := 10;
       ELSIF (#tempOffTime.DAY > 9)
       THEN
         #tempOffTime.DAY := 9;
       END_IF;

       IF (#tempActTime >= #tempOnTime)
         AND (#tempActTime < #tempOffTime)
       THEN
         #tempSignal := true;
       ELSE
         #tempSignal := false;
       END_IF;

       #signal := #tempSignal;

     6:  // Mode: weekend (Saturday and Sunday)    
       #tempOnTime.YEAR := 2015;
       #tempOnTime.MONTH := 1;
       #tempOnTime.DAY := #tempTime.WEEKDAY + 3;

       IF (#tempOnTime.DAY < 10)
       THEN
         #tempOnTime := #tempOnTime + t#7d;
       END_IF;

       #tempOnTimeTOD := DTL_TO_TOD(#tempOnTime);

       #tempOffTime.YEAR := 2015;
       #tempOffTime.MONTH := 1;
       #tempOffTime.DAY := #tempTime.WEEKDAY + 3;

       IF (#tempOffTime.DAY < 10)
       THEN
         #tempOffTime := #tempOffTime + t#7d;
       END_IF;

       #tempOffTimeTOD := DTL_TO_TOD(#tempOffTime);

       #tempActTime := #tempTime;
       #tempActTime.YEAR := 2015;
       #tempActTime.MONTH := 1;
       #tempActTime.DAY := #tempActTime.WEEKDAY + 3;

       IF (#tempActTime.DAY < 10)
       THEN
         #tempActTime := #tempActTime + t#7d;
       END_IF;

       #tempActTimeTOD := DTL_TO_TOD(#tempTime);

       IF (#tempOnTimeTOD > #tempOffTimeTOD)
       THEN
         #tempCrossMidnight := TRUE;
         IF (#tempActTimeTOD > #tempOffTimeTOD)
         THEN
           #tempOffTime := #tempOffTime + t#1d;
         ELSE
           #tempOnTime := #tempOnTime - t#1d;
         END_IF;
       ELSE
         #tempCrossMidnight := FALSE;
       END_IF;

       IF (#tempOnTime.DAY < 10)
       THEN
         #tempOnTime.DAY := 10;
       ELSIF (#tempOnTime.DAY > 11)
       THEN
         #tempOnTime.DAY := 11;
       END_IF;

       IF (#tempOffTime.DAY > 11)
         AND (#tempCrossMidnight = TRUE)
       THEN
         #tempOffTime.DAY := 12;
       ELSIF (#tempOffTime.DAY > 11)
       THEN
         #tempOffTime.DAY := 11;
       END_IF;

       IF (#tempActTime >= #tempOnTime)
         AND (#tempActTime < #tempOffTime)
       THEN
         #tempSignal := true;
       ELSE
         #tempSignal := false;
       END_IF;

       #signal := #tempSignal;

     ELSE
       #error := true;
       #statusID := #ERROR_IN_THIS_BLOCK;
       #status := #NO_MODE_SELECTED;
       RETURN;
   END_CASE;